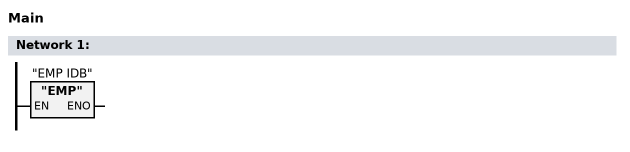
   RUNG wire#powerrail
      "EMP IDB"()
   END_RUNG
   // the same network as SCL:
   "EMP IDB"();   // "EMP"
END_REGION
END_ORGANIZATION_BLOCK

// folder: Display: LED

FUNCTION_BLOCK "LED_Request_Table"   // FB60, SCL
{ S7_Optimized_Access := 'TRUE' }
VERSION : 0.1
   VAR_INPUT
      pn_library : "Recipe: PN Text Library";
      saved_wips : "Recipe: HMI Stations Saved Wips";
      stations : "Station: All Stations";
      table_data : "Part Request Data";
   END_VAR
   VAR_IN_OUT
      request_table : "LED Sign Data";
   END_VAR
   VAR
      row_indices : Array[0..11] of DInt;
   END_VAR
   // row_indices[0] := 0;
   // row_indices[1] := 1;
   // row_indices[2] := 2;
   // row_indices[3] := 3;
   // row_indices[4] := 4;
   // row_indices[5] := 5;
   // row_indices[6] := 6;
   // row_indices[7] := 7;
   // row_indices[8] := 8;
   // row_indices[9] := 9;
   // row_indices[10] := 10;
   // row_indices[11] := 11;
BEGIN
   "Request_Table.Draw"(pn_library := #pn_library,
                        row_indices := #row_indices,
                        saved_wips := #saved_wips,
                        stations := #stations,
                        table_data := #table_data,
                        request_table := #request_table.row);
END_FUNCTION_BLOCK

// folder: Display: Warehouse/001 Request Table

FUNCTION_BLOCK "HMI_Request_Table"   // FB16, SCL
{ S7_Optimized_Access := 'TRUE' }
VERSION : 0.1
   VAR_INPUT
      pn_library : "Recipe: PN Text Library";
      saved_wips : "Recipe: HMI Stations Saved Wips";
      stations : "Station: All Stations";
      table_data : "Part Request Data";
   END_VAR
   VAR_IN_OUT
      barcode_data : "Barcode.UDT";
      request_table : "Part Call Screen";
      request_table_navigation : "Nav Bar Data: PLC";
   END_VAR
   VAR RETAIN
      row_indices : Array[0.."PART_REQUEST_ROW_COUNT_WAREHOUSE_HMI"] of DInt;
   END_VAR
   VAR
      Table_Navigation : "Table Nav";
      Row_Selection : "Request_Table.Row_Selection";
   END_VAR
   // row_indices[1] := 1;
   // row_indices[2] := 2;
   // row_indices[3] := 3;
   // row_indices[4] := 4;
   // row_indices[5] := 5;
   // row_indices[6] := 6;
   // row_indices[7] := 7;
   // row_indices[8] := 8;
   // row_indices[9] := 9;
   // row_indices[10] := 10;
BEGIN
   REGION "TABLE NAVIGATION"
       #Table_Navigation(tblData := #table_data.row,
                         tblDisp := #request_table.row,
                         tableNav := #request_table_navigation,
                         rowIndices := #row_indices);
   END_REGION


   REGION "NAV BUTTON ANIMATIONS"
       "Request_Table.Navigation_Animations"(#request_table_navigation);
   END_REGION


   REGION "DRAW TABLE"
       "Request_Table.Draw"(pn_library := #pn_library,
                            row_indices := #row_indices,
                            saved_wips := #saved_wips,
                            stations := #stations,
                            table_data := #table_data,
                            request_table := #request_table.row);
   END_REGION


   REGION "LOAD SELECTION DATA"
       #Row_Selection(request_table := #request_table,
                      barcode_data := #barcode_data);
   END_REGION
END_FUNCTION_BLOCK

FUNCTION "Address in Loaded Wip" : Bool   // FC43, SCL
{ S7_Optimized_Access := 'TRUE' }
VERSION : 0.1
   VAR_INPUT
      pWip : DInt;
      stn : "Station: Single Station";
   END_VAR
   VAR_TEMP
      ret : Bool;
   END_VAR
BEGIN
   IF #pWip = #stn.wipData.index THEN
       #ret := TRUE;
   END_IF;
   #"Address in Loaded Wip" := #ret;
END_FUNCTION

// folder: Display: Warehouse/002 Settings

FUNCTION_BLOCK "Settings Screen"   // FB19, SCL
{ S7_Optimized_Access := 'TRUE' }
VERSION : 0.1
   VAR_INPUT
      settings_meta : "Setting Meta Data";
      wip_library : "Recipe: Wip Text Library";
   END_VAR
   VAR_IN_OUT
      pn_library : "Recipe: PN Text Library";
      saved_wips : "Recipe: HMI Stations Saved Wips";
      stations : "Station: All Stations";
      settings : "Settings";
   END_VAR
   VAR
      "Assign Button" : "Assign Button";
      "Critical Time IO Field" : "Critical_IO_Field";
      "Dropzone IO Field" : "Dropzone_IO_Field";
      first_row : DInt;
      "Line IO Field" : "Line_IO_Field";
      "Part Number IO Field" : "Part Number IO Field";
      processed_inputs : "Settings Screen: Processed Inputs";
      "Select Buttons Button" : "Select Buttons";
      "Select Station Button" : "Select Station PB";
      "Select WIP Button" : "Select WIP PB";
      "Table Nav_Instance" : "Table Nav";
      "Total Time IO Field" : "Total_IO_Field";
      "WIP Select Table NavBar" : "NavBar";
      inst_Selected_WIP_Table : "Selected_WIP_Table";
   END_VAR
   VAR_TEMP
      _station_rows_buffer : Array[0..2] of "Settings Station Row Data";
   END_VAR
   VAR CONSTANT
      TABLE_LENGTH : DInt := 49;
      VISIBLE_ROW_COUNT : DInt := 2;
   END_VAR
BEGIN
   REGION "SELECT STATION BUTTON"
       #"Select Station Button"(#settings.selectStation);
   END_REGION

   REGION "SELECT BUTTONS BUTTON"
       #"Select Buttons Button"(settings_meta := #settings_meta,
                                stations := #stations,
                                interface := #settings.selectButton);
   END_REGION

   REGION "SELECT WIP BUTTON"
       #"Select WIP Button"(settings_meta := #settings_meta,
                            stations := #stations,
                            interface := #settings.selectWip);
   END_REGION

   REGION "LINE IO FIELD"
       #"Line IO Field"(settings_meta := #settings_meta,
                        stations := #stations,
                        interface := #settings.line,
                        get_line := #processed_inputs.line_name);
   END_REGION

   REGION "DROPZONE IO FIELD"
       #"Dropzone IO Field"(settings_meta := #settings_meta,
                            stations := #stations,
                            interface := #settings.dropzone,
                            get_dropzone := #processed_inputs.dropzone);
   END_REGION

   REGION "TOTAL TIME IO FIELD"
       #"Total Time IO Field"(settings_meta := #settings_meta,
                              stations := #stations,
                              interface := #settings.total,
                              state_changes := #processed_inputs.total);
   END_REGION

   REGION "CRITICAL TIME IO FIELD"
       #"Critical Time IO Field"(settings_meta := #settings_meta,
                                 stations := #stations,
                                 interface := #settings.critical,
                                 state_changes := #processed_inputs.critical);
   END_REGION

   REGION "PART NUMBER ENTRY FIELD"
       #"Part Number IO Field"(settings_meta := #settings_meta,
                               stations := #stations,
                               part_number_library := #pn_library,
                               interface := #settings.partNumber,
                               processed_part_number_entry := #processed_inputs.part_number);

   END_REGION

   REGION "ASSIGN BUTTON"
       #"Assign Button"(processed_inputs := #processed_inputs,
                        settings := #settings,
                        settings_meta := #settings_meta,
                        pn_library := #pn_library,
                        saved_wips := #saved_wips,
                        stations := #stations,
                        interface := #settings.assign,
                        state_changes := #processed_inputs.assign);
   END_REGION

   REGION "SELECTED WIP TABLE"
       #_station_rows_buffer := #settings.stationRows;
       #inst_Selected_WIP_Table(saved_wips := #saved_wips,
                                settings_meta := #settings_meta,
                                stations := #stations,
                                wip_library := #wip_library,
                                pn_library := #pn_library,
                                navigation_bar := #settings.stnTableNavBar.plc,
                                stationRows := #_station_rows_buffer);
       #settings.stationRows := #_station_rows_buffer;
   END_REGION

   REGION "WIP SELECT TABLE NAVBAR"
       #"WIP Select Table NavBar"(hide := #settings_meta.selected_stations.count < 4,
                                  TABLE_LENGTH := #TABLE_LENGTH,
                                  VISIBLE_ROW_COUNT := #VISIBLE_ROW_COUNT,
                                  interface := #settings.stnTableNavBar,
                                  first_row := #first_row);
   END_REGION
END_FUNCTION_BLOCK

FUNCTION "Settings Screen: Load Selected: Non-HMI Station" : Void   // FC150, SCL
{ S7_Optimized_Access := 'TRUE' }
VERSION : 0.1
   VAR_INPUT
      stations : "Station: All Stations";
      selected_stations : "Selected Stations";
      wip_library : "Recipe: Wip Text Library";
      part_number_library : "Recipe: PN Text Library";
   END_VAR
   VAR_IN_OUT
      selected_station_table : Array[0..2] of "Settings Station Row Data";
   END_VAR
   VAR_TEMP
      station_index : Int;
      table_row_index : Int;
   END_VAR
BEGIN
   FOR #station_index := 0 TO "STATION_COUNT" DO
       IF #selected_stations.stns[#station_index] THEN
           "Settings Screen: Load Selected WIP"(station := #stations.stn[#station_index],
                                                wip_library := #wip_library,
                                                part_number_library := #part_number_library,
                                                table_row := #selected_station_table[#table_row_index]);
           #table_row_index += 1;
           IF #table_row_index > 2 THEN
               EXIT;
           END_IF;
       END_IF;
   END_FOR;
END_FUNCTION

FUNCTION "Settings Screen: Load Selected WIP" : Void   // FC151, SCL
{ S7_Optimized_Access := 'TRUE' }
VERSION : 0.1
   VAR_INPUT
      station : "Station: Single Station";
      wip_library : "Recipe: Wip Text Library";
      part_number_library : "Recipe: PN Text Library";
   END_VAR
   VAR_IN_OUT
      table_row : "Settings Station Row Data";
   END_VAR
   VAR_TEMP
      _table_row : "Settings Station Row Data";
      button_index : Int;
   END_VAR
BEGIN
   REGION "NOTES"
       (*
       Simple data map from station presented at input to hmi data structure.
       Decision about which data to map is done in parent.
       last edit: 2021-10-06
       *)
   END_REGION

   REGION "BUFFER IN"
       #_table_row := #table_row;
   END_REGION

   REGION "MAP"
       #_table_row.line.data := #station.id.lineName;
       #_table_row.dropzone.data := "Strip Sign"(USINT_TO_WSTRING(#station.id.dropZone));
       #_table_row.wip.data := "WIP.Code_to_WString"(wipTxtLib := #wip_library,
                                                           code := #station.wipData.code);
       FOR #button_index := 0 TO "BUTTON_COUNT" DO
           "Settings Screen: Load Selected WIP: Load Button"(wip_components:=#station.wipCmpts,
                                                                 wip_library := #wip_library,
                                                                 button_index := #button_index,
                                                                 part_number_liberary := #part_number_library,
                                                                 button_row := #_table_row.btnRows[#button_index]);
       END_FOR;
   END_REGION

   REGION "BUFFER OUT"
       #table_row := #_table_row;
   END_REGION
END_FUNCTION

FUNCTION "Settings Screen: Selected Station Table Row Color" : Void   // FC152, SCL
{ S7_Optimized_Access := 'TRUE' }
VERSION : 0.1
BEGIN
END_FUNCTION

FUNCTION "Settings Screen: Load Selected WIP: Load Button" : Void   // FC155, SCL
{ S7_Optimized_Access := 'TRUE' }
VERSION : 0.1
   VAR_INPUT
      button_index : Int;
      part_number_liberary : "Recipe: PN Text Library";
      wip_components : "Station: Wip: Wip Module";
      wip_library : "Recipe: Wip Text Library";
   END_VAR
   VAR_IN_OUT
      button_row : "Settings Station Row Button Row Data";
   END_VAR
   VAR_TEMP
      _button_row : "Settings Station Row Button Row Data";
      part_number_wstring : WString;
      part_number_code : DInt;
   END_VAR
   VAR CONSTANT
      no_code : WString;
   END_VAR
BEGIN
   REGION "NOTES"
       (*
       Simple data map from station presented at input to hmi data structure.
       Decision about which data to map is done in parent.
       last edit: 2021-10-06
       *)
   END_REGION

   REGION "BUFFER IN"    
       #_button_row := #button_row;
   END_REGION

   REGION "BUTTON LABEL"
       // CURRENTLY A STATIC LABEL
   END_REGION

   REGION "ALOTTED TIME"
       #_button_row.total.data := "Timer.Real_to_WString"(#wip_components.timers.ptAllotted[#button_index]);
   END_REGION

   REGION "CRITICAL TIME"
       #_button_row.critical.data := "Timer.Real_to_WString"(#wip_components.timers.ptCritical[#button_index]);
   END_REGION

   REGION "PART NUMBER"

       REGION "PROCESS PART NUMBER"
           #part_number_code := #wip_components.pnCode[#button_index];
           #part_number_wstring := "Part_Number.Code_to_WString"(pnLib := #part_number_liberary,
                                                         pnCode := #part_number_code);
       END_REGION

       REGION "SINGLE LINE PART NUMBER"
           IF "Part_Number.Is_Single"(#part_number_code) THEN
               #_button_row.singlePN.data := #part_number_wstring;
               #_button_row.doublePN.data := #no_code;
           END_IF;
       END_REGION

       REGION "DOUBLE LINE PART NUMBER"
           IF "Part_Number.Is_Double"(#part_number_code) THEN
               #_button_row.singlePN.data := #no_code;
               #_button_row.doublePN.data := #part_number_wstring;
           END_IF;
       END_REGION

   END_REGION

   REGION "BUFFER OUT"
       #button_row := #_button_row;
   END_REGION
END_FUNCTION

FUNCTION "Settings Screen: Load Selected: HMI Station" : Void   // FC176, SCL
{ S7_Optimized_Access := 'TRUE' }
VERSION : 0.1
   VAR_INPUT
      stations : "Station: All Stations";
      selected_wips : "Selected Wips";
      wip_library : "Recipe: Wip Text Library";
      part_number_library : "Recipe: PN Text Library";
   END_VAR
   VAR_IN_OUT
      selected_station_table : Array[0..2] of "Settings Station Row Data";
   END_VAR
   VAR_TEMP
      station_index : Int;
      table_row_index : Int;
   END_VAR
BEGIN
   FOR #station_index := 0 TO #selected_wips.count DO
       "Settings Screen: Load Selected WIP"(station := #stations.stn[#station_index],
                                            wip_library := #wip_library,
                                            part_number_library := #part_number_library,
                                            table_row := #selected_station_table[#table_row_index]);END_FOR;
END_FUNCTION

// folder: Display: Warehouse/002 Settings/Assign Button

FUNCTION_BLOCK "Assign Button"   // FB55, SCL
{ S7_Optimized_Access := 'TRUE' }
VERSION : 0.1
   VAR_INPUT
      processed_inputs : "Settings Screen: Processed Inputs";
      settings : "Settings";
      settings_meta : "Setting Meta Data";
   END_VAR
   VAR_IN_OUT
      interface : "Push Button Data";
      pn_library : "Recipe: PN Text Library";
      saved_wips : "Recipe: HMI Stations Saved Wips";
      state_changes : "Push Button Data: State Change Data";
      stations : "Station: All Stations";
   END_VAR
   VAR
      "Push Button: State Changes" : "Push Button: State Changes";
   END_VAR
   VAR_TEMP
      _interface : "Push Button Data";
      _state_changes : "Push Button Data: State Change Data";
   END_VAR
BEGIN
   REGION "BUFFER IN"
       #_interface := #interface;
   END_REGION


   REGION "PROCESS USER INPUT"
       #"Push Button: State Changes"(interface := #_interface,
                                     state_changes := #_state_changes);
   END_REGION


   REGION "ANIMATE"
       "Assign_Button.Animate"(settings_meta := #settings_meta,
                                         interface := #_interface);
   END_REGION


   REGION "PERFOM ASSIGNMNET"
       IF #_state_changes.actuate.falling THEN
           "Assign_Button.Perform_Assignment"(processed_inputs := #processed_inputs,
                                              settings := #settings,
                                              settings_meta := #settings_meta,
                                              pn_library := #pn_library,
                                              stations := #stations,
                                              saved_wips := #saved_wips);
       END_IF;
   END_REGION


   REGION "BUFFER OUT"
       #interface := #_interface;
       #state_changes := #_state_changes;
   END_REGION
END_FUNCTION_BLOCK

FUNCTION "Assign_Button.Make_Visible_Enable" : Bool   // FC197, SCL
{ S7_Optimized_Access := 'TRUE' }
VERSION : 0.1
   VAR_INPUT
      setting_meta : "Setting Meta Data";
   END_VAR
BEGIN
   #"Assign_Button.Make_Visible_Enable" :=  #setting_meta.selected_btns.count > 0;
END_FUNCTION

FUNCTION "Assign_Button.Animate" : Void   // FC198, SCL
{ S7_Optimized_Access := 'TRUE' }
VERSION : 0.1
   VAR_INPUT
      settings_meta : "Setting Meta Data";
   END_VAR
   VAR_IN_OUT
      interface : "Push Button Data";
   END_VAR
   VAR_TEMP
      selected_station_count : DInt;
   END_VAR
BEGIN
   REGION "COLOR"
   #interface.animate := "WHITE_BACKGROUND";
   END_REGION

   REGION "VISIBILITY
       #interface.visible := "Assign_Button.Make_Visible_Enable"(setting_meta := #settings_meta);
   END_REGION

   REGION "ENABLE"
       #interface.enable := "Assign_Button.Make_Visible_Enable"(setting_meta := #settings_meta);
   END_REGION
END_FUNCTION

FUNCTION "Assign_Button.Perform_Assignment" : Void   // FC235, SCL
{ S7_Optimized_Access := 'TRUE' }
VERSION : 0.1
   VAR_INPUT
      processed_inputs : "Settings Screen: Processed Inputs";
      settings : "Settings";
      settings_meta : "Setting Meta Data";
   END_VAR
   VAR_IN_OUT
      pn_library : "Recipe: PN Text Library";
      stations : "Station: All Stations";
      saved_wips : "Recipe: HMI Stations Saved Wips";
   END_VAR
   VAR_TEMP
      _station_indices : Array[0.."STATION_COUNT"] of Int;
   END_VAR
BEGIN
   REGION "DO NOTHING ON NO SELECTED STAION"
       IF #settings_meta.selected_stations.count = 0 THEN
           RETURN;
       END_IF;
   END_REGION


   REGION "HMI STATIONS"
       "Selected_Stations.Indices"(selected_stations:=#settings_meta.selected_stations,
                                   selected_stations_indices:=#_station_indices);
       IF "Is_HMI_Station"(#stations.stn[#_station_indices[0]]) THEN
           "Assign_Button.HMI_Stations"(processed_inputs := #processed_inputs,
                                        settings := #settings,
                                        settings_meta := #settings_meta,
                                        pn_library := #pn_library,
                                        saved_wips := #saved_wips,
                                        stations := #stations);
           RETURN;
       END_IF;
   END_REGION


   REGION "KP8 STATIONS"
       "Assign_Button.KP8_Station"(processed_inputs := #processed_inputs,
                                   settings := #settings,
                                   settings_meta := #settings_meta,
                                   all_stations := #stations,
                                   pn_library := #pn_library);
       RETURN;
   END_REGION
END_FUNCTION

FUNCTION "Assign_Button.Assign_ID_Parameters" : Void   // FC264, SCL
{ S7_Optimized_Access := 'TRUE' }
VERSION : 0.1
   VAR_INPUT
      processed_inputs : "Settings Screen: Processed Inputs";
      settings : "Settings";
   END_VAR
   VAR_IN_OUT
      id : "Station: Id";
   END_VAR
BEGIN
   IF #settings.line.enable THEN
       #id.lineName := #processed_inputs.line_name.actual;
   END_IF;
   IF #settings.dropzone.enable THEN
       #id.dropZone := #processed_inputs.dropzone.actual;
   END_IF;
END_FUNCTION

// folder: Display: Warehouse/002 Settings/Assign Button/HMI Station

FUNCTION "Assign_Button.HMI_Stations" : Void   // FC236, SCL
{ S7_Optimized_Access := 'TRUE' }
VERSION : 0.1
   VAR_INPUT
      processed_inputs : "Settings Screen: Processed Inputs";
      settings : "Settings";
      settings_meta : "Setting Meta Data";
   END_VAR
   VAR_IN_OUT
      pn_library : "Recipe: PN Text Library";
      saved_wips : "Recipe: HMI Stations Saved Wips";
      stations : "Station: All Stations";
   END_VAR
   VAR_TEMP
      _i : Int;
      _length : Int;
      _selected_stations : Array[0.."STATION_COUNT"] of Int;
      _p_station : Int;
   END_VAR
BEGIN
   REGION "DO NOTHING IF NO STATIONS SELECTED"
       IF #settings_meta.selected_stations.count = 0 THEN
           RETURN;
       END_IF;
   END_REGION


   REGION "GET INDICES OF SELECTED STATIONS"
       "Selected_Stations.Indices"(selected_stations := #settings_meta.selected_stations,
                                   selected_stations_indices := #_selected_stations);

   END_REGION


   REGION "FOR EACH SELECTED STATION"
       #_length := UDINT_TO_INT("Array.Any.Length"(#saved_wips.stn)) - 1;
       FOR #_i := 0 TO #_length DO

           IF #_selected_stations[#_i] = "NULL_TOKEN" THEN
               RETURN;
           END_IF;

           REGION "ASSIGN TO WIP"
               "Assign_Button.Assign_ID_Parameters"(processed_inputs := #processed_inputs,
                                                    settings := #settings,
                                                    id := #stations.stn[#_selected_stations[#_i]].id);
               #_p_station := "WIP.Global_Index_to_HMI_Station_Index"(global_index := #_selected_stations[#_i],
                                                                      saved_WIPs := #saved_wips);
               "Assign_Button.HMI_Stations.WIP"(processed_inputs:=#processed_inputs,
                                                selected_wips := #settings_meta.selected_wips,
                                                selected_buttons := #settings_meta.selected_btns,
                                                pn_library := #pn_library,
                                                stations_wips := #saved_wips.stn[#_p_station]);
           END_REGION

       END_FOR;
   END_REGION
END_FUNCTION

FUNCTION "Assign_Button.HMI_Stations.WIP" : Void   // FC237, SCL
{ S7_Optimized_Access := 'TRUE' }
VERSION : 0.1
   VAR_INPUT
      processed_inputs : "Settings Screen: Processed Inputs";
      selected_wips : "Selected Wips";
      selected_buttons : "Selected Buttons";
   END_VAR
   VAR_IN_OUT
      pn_library : "Recipe: PN Text Library";
      stations_wips : "WIP: Station";
   END_VAR
   VAR_TEMP
      _i : Int;
      _p_wip : Int;
      _selected_wip_indices : Array[0.."WIP_COUNT"] of Int;
   END_VAR
BEGIN
   REGION "DO NOTHING IF NO WIPS SELECTED"
       IF #selected_wips.count = 0 THEN
           RETURN;
       END_IF;
   END_REGION


   REGION "GET INDICES OF SELECTED WIPS"    
       "WIP_Station.Indices_of_Selected_WIPs"(selected_wips := #selected_wips,
                                              station_wips := #stations_wips,
                                              selected_wip_indices := #_selected_wip_indices);
   END_REGION


   REGION "FOR EACH SELECTED WIP"
       FOR #_i := 0 TO #selected_wips.count DO

           REGION "ASSIGN DATA TO SELECTED BUTTONS"
               #_p_wip := #_selected_wip_indices[#_i];
               IF #_p_wip = "NULL_TOKEN" THEN
                   RETURN;
               END_IF;
               "Assign_Button.HMI_Stations.WIP.Buttons"(processed_inputs := #processed_inputs,
                                                        selected_buttons := #selected_buttons,
                                                        pn_library := #pn_library,
                                                        wip_module := #stations_wips.wip[#_p_wip]);
           END_REGION

       END_FOR;
   END_REGION
END_FUNCTION

FUNCTION "Assign_Button.HMI_Stations.WIP.Buttons" : Void   // FC238, SCL
{ S7_Optimized_Access := 'TRUE' }
VERSION : 0.1
   VAR_INPUT
      processed_inputs : "Settings Screen: Processed Inputs";
      selected_buttons : "Selected Buttons";
   END_VAR
   VAR_IN_OUT
      pn_library : "Recipe: PN Text Library";
      wip_module : "Station: Wip: Wip Module";
   END_VAR
   VAR_TEMP
      _i : Int;
      _p_btn : Int;
      _selected_buttons_indices : Array[0..7] of Int;
   END_VAR
BEGIN
   REGION "DO NOTHING IF NO BUTTONS SELECTED
       IF #selected_buttons.count = 0 THEN
           RETURN;
       END_IF;
   END_REGION


   REGION "GET INDICES OF SELECTED BUTTONS"
       "Selected_Buttons.Indices"(selected_buttons := #selected_buttons,
                                  selected_buttons_indices := #_selected_buttons_indices);
   END_REGION

   REGION "FOR EACH SELECTED BUTTON"
       FOR #_i := 0 TO #selected_buttons.count DO

           REGION "ASSIGN DATA TO SELECTED BUTTON"
               #_p_btn := #_selected_buttons_indices[#_i];
               "Assign_Button.HMI_Stations.Assign_Station_Button_Data"(processed_inputs := #processed_inputs,
                                                                       index := #_p_btn,
                                                                       pn_library := #pn_library,
                                                                       wip_module := #wip_module);
           END_REGION

       END_FOR;
   END_REGION
END_FUNCTION

FUNCTION "Assign_Button.HMI_Stations.Assign_Station_Button_Data" : Void   // FC239, SCL
{ S7_Optimized_Access := 'TRUE' }
VERSION : 0.1
   VAR_INPUT
      processed_inputs : "Settings Screen: Processed Inputs";
      index : Int;
   END_VAR
   VAR_IN_OUT
      pn_library : "Recipe: PN Text Library";
      wip_module : "Station: Wip: Wip Module";
   END_VAR
BEGIN
   IF #index = "NULL_TOKEN" THEN
       RETURN;
   END_IF;
   #wip_module.pnCode[#index] := "Part_Number.WString_to_Code"(part_number := #processed_inputs.part_number.actual,
                                                               pn_library := #pn_library);
   #wip_module.timers.ptAllotted[#index] := #processed_inputs.total.actual;
   #wip_module.timers.ptCritical[#index] := #processed_inputs.critical.actual;
END_FUNCTION

// folder: Display: Warehouse/002 Settings/Assign Button/KP8 Station

FUNCTION "Assign_Button.KP8_Station" : Void   // FC247, SCL
{ S7_Optimized_Access := 'TRUE' }
VERSION : 0.1
   VAR_INPUT
      processed_inputs : "Settings Screen: Processed Inputs";
      settings : "Settings";
      settings_meta : "Setting Meta Data";
   END_VAR
   VAR_IN_OUT
      all_stations : "Station: All Stations";
      pn_library : "Recipe: PN Text Library";
   END_VAR
   VAR_TEMP
      _i : Int;
      _length : Int;
      _selected_stations : Array[0.."STATION_COUNT"] of Int;
      _p_station : Int;
   END_VAR
BEGIN
   REGION "DO NOTHING IF NO STATIONS SELECTED"
       IF #settings_meta.selected_stations.count = 0 THEN
           RETURN;
       END_IF;
   END_REGION


   REGION "GET INDICES OF SELECTED STATIONS"
       "Selected_Stations.Indices"(selected_stations := #settings_meta.selected_stations,
                                   selected_stations_indices := #_selected_stations);
   END_REGION


   REGION "FOR EACH SELECTED STATION"
       IF #settings_meta.selectable_stations.count = 0 THEN
           RETURN;
       END_IF;
       FOR #_i := 0 TO #settings_meta.selected_stations.count DO
           IF #_selected_stations[#_i] = "NULL_TOKEN" THEN
               RETURN;
           END_IF;
           #_p_station := #_selected_stations[#_i];
           "Assign_Button.Assign_ID_Parameters"(processed_inputs := #processed_inputs,
                                                settings := #settings,
                                                id := #all_stations.stn[#_p_station].id);
           "Assign_Button.KP8_Stations.Buttons"(processed_inputs := #processed_inputs,
                                                selected_buttons := #settings_meta.selected_btns,
                                                pn_library := #pn_library,
                                                station := #all_stations.stn[#_p_station]);
       END_FOR;
   END_REGION
END_FUNCTION

FUNCTION "Assign_Button.KP8_Station.Assign_Station_Button_Data" : Void   // FC248, SCL
{ S7_Optimized_Access := 'TRUE' }
VERSION : 0.1
   VAR_INPUT
      button_number : Int;
      processed_inputs : "Settings Screen: Processed Inputs";
   END_VAR
   VAR_IN_OUT
      pn_library : "Recipe: PN Text Library";
      station : "Station: Single Station";
   END_VAR
   VAR_TEMP
      _i : Int;
      _length : Int;
      _selected_stations : Array[0.."STATION_COUNT"] of Int;
      _p_station : Int;
   END_VAR
BEGIN
   IF #button_number = "NULL_TOKEN" THEN
       RETURN;
   END_IF;
   #station.wipCmpts.pnCode[#button_number] := "Part_Number.WString_to_Code"(part_number := #processed_inputs.part_number.actual,
                                                                             pn_library := #pn_library);
   #station.wipCmpts.timers.ptCritical[#button_number] := #processed_inputs.critical.actual;
   #station.wipCmpts.timers.ptAllotted[#button_number] := #processed_inputs.total.actual;
END_FUNCTION

FUNCTION "Assign_Button.KP8_Stations.Buttons" : Void   // FC249, SCL
{ S7_Optimized_Access := 'TRUE' }
VERSION : 0.1
   VAR_INPUT
      processed_inputs : "Settings Screen: Processed Inputs";
      selected_buttons : "Selected Buttons";
   END_VAR
   VAR_IN_OUT
      pn_library : "Recipe: PN Text Library";
      station : "Station: Single Station";
   END_VAR
   VAR_TEMP
      _i : Int;
      _p_btn : Int;
      _selected_buttons_indices : Array[0..7] of Int;
   END_VAR
BEGIN
   REGION "DO NOTHING IF NO BUTTONS SELECTED
       IF #selected_buttons.count = 0 THEN
           RETURN;
       END_IF;
   END_REGION


   REGION "GET INDICES OF SELECTED BUTTONS"
       "Selected_Buttons.Indices"(selected_buttons := #selected_buttons,
                                  selected_buttons_indices := #_selected_buttons_indices);
   END_REGION


   REGION "FOR EACH SELECTED BUTTON"
       FOR #_i := 0 TO #selected_buttons.count - 1 DO

           IF #_selected_buttons_indices[#_i] = "NULL_TOKEN" THEN
               RETURN;
           END_IF;

           REGION "ASSIGN DATA TO SELECTED BUTTON"
               #_p_btn := #_selected_buttons_indices[#_i];
               "Assign_Button.KP8_Station.Assign_Station_Button_Data"(button_number := #_p_btn,
                                                                      processed_inputs := #processed_inputs,
                                                                      pn_library := #pn_library,
                                                                      station := #station);
           END_REGION

       END_FOR;
   END_REGION
END_FUNCTION

// folder: Display: Warehouse/002 Settings/Critical IO Field

FUNCTION_BLOCK "Critical_IO_Field"   // FB53, SCL
{ S7_Optimized_Access := 'TRUE' }
VERSION : 0.1
   VAR_INPUT
      settings_meta : "Setting Meta Data";
      stations : "Station: All Stations";
   END_VAR
   VAR_IN_OUT
      interface : "IO Field Data: Label with Data";
      state_changes : "State Changes: Real";
   END_VAR
   VAR
      Critical_IO_Field : "IO Field: State Changes";
      Detect_Stat_Changes : "Real.State_Change";
   END_VAR
   VAR_TEMP
      _interface : "IO Field Data: Label with Data";
      feedback : "IO Field: State Change Data";
   END_VAR
BEGIN
   REGION "BUFFER IN"
       #_interface := #interface;
   END_REGION

   REGION "PROCESS USER INPUT"
       #Critical_IO_Field(interface := #_interface,
                          feedback := #feedback);
       #Detect_Stat_Changes(value := "Timer.WString_to_Real"(#_interface.value),
                            get_real := #state_changes);
   END_REGION

   REGION "BUFFER OUT"
       "Critical_IO_Field.Animate"(feedback := #feedback,
                                   settings_meta := #settings_meta,
                                   stations := #stations,
                                   interface := #_interface);
   END_REGION

   REGION "BUFFER OUT"
       #interface := #_interface;
   END_REGION
END_FUNCTION_BLOCK

FUNCTION "Critical_IO_Field.Make_Visible_Enable" : Bool   // FC191, SCL
{ S7_Optimized_Access := 'TRUE' }
VERSION : 0.1
   VAR_INPUT
      setting_meta : "Setting Meta Data";
   END_VAR
BEGIN
   #"Critical_IO_Field.Make_Visible_Enable" :=  #setting_meta.selected_btns.count > 0;
END_FUNCTION

FUNCTION "Critical_IO_Field.Animate" : Void   // FC192, SCL
{ S7_Optimized_Access := 'TRUE' }
VERSION : 0.1
   VAR_INPUT
      feedback : "IO Field: State Change Data";
      settings_meta : "Setting Meta Data";
      stations : "Station: All Stations";
   END_VAR
   VAR_IN_OUT
      interface : "IO Field Data: Label with Data";
   END_VAR
   VAR_TEMP
      _visible_enabled : Bool;
   END_VAR
BEGIN
   REGION "COLOR"
   #interface.animate := "WHITE_BACKGROUND";
   END_REGION


   REGION "SET STATE"
       #_visible_enabled := "Critical_IO_Field.Make_Visible_Enable"(setting_meta := #settings_meta);
   END_REGION


   REGION "VISIBILITY
       #interface.visible := #_visible_enabled;
   END_REGION


   REGION "ENABLE"
       #interface.enable := #_visible_enabled;
   END_REGION


   REGION "POPULATE VALUE"
       IF #settings_meta.button_selection_change.selection_change THEN
           #interface.value := "Critical_IO_Field.Populate_Value"(hidden := NOT #_visible_enabled,
                                                                  selected_buttons := #settings_meta.selected_btns,
                                                                  selected_stations := #settings_meta.selected_stations,
                                                                  stations := #stations);
       END_IF;
   END_REGION
END_FUNCTION

FUNCTION "Critical_IO_Field.Populate_Value" : WString   // FC283, SCL
{ S7_Optimized_Access := 'TRUE' }
VERSION : 0.1
   VAR_INPUT
      hidden : Bool;
      selected_buttons : "Selected Buttons";
      selected_stations : "Selected Stations";
      stations : "Station: All Stations";
   END_VAR
   VAR_TEMP
      _critical : WString;
      _p_station : Int;
      _p_button : Int;
   END_VAR
   VAR CONSTANT
      BLANK : WString;
      ZERO : WChar := WCHAR#'0';
   END_VAR
BEGIN
   IF #hidden THEN
       #"Critical_IO_Field.Populate_Value" := #BLANK;
       RETURN;
   END_IF;
   #_p_station := "Selected_Stations.Get_First_Selected_Station"(#selected_stations);
   #_p_button := "Selected_Buttons.Get_First_Selected_Button"(#selected_buttons);
   #_critical := "Timer.Real_to_WString"(#stations.stn[#_p_station].wipCmpts.timers.ptCritical[#_p_button]);
   #"Critical_IO_Field.Populate_Value" := #_critical;
END_FUNCTION

// folder: Display: Warehouse/002 Settings/Dropzone IO Field

FUNCTION_BLOCK "Dropzone_IO_Field"   // FB50, SCL
{ S7_Optimized_Access := 'TRUE' }
VERSION : 0.1
   VAR_INPUT
      settings_meta : "Setting Meta Data";
      stations : "Station: All Stations";
   END_VAR
   VAR_IN_OUT
      interface : "IO Field Data: Label with Data";
      get_dropzone : "State Changes: USInt";
   END_VAR
   VAR
      "Line IO Field" : "IO Field: State Changes";
      "Get Dropzone Input" : "USInt.State_change";
   END_VAR
   VAR_TEMP
      _feedback : "IO Field: State Change Data";
      _interface : "IO Field Data: Label with Data";
   END_VAR
BEGIN
   REGION "BUFFER IN"
       #_interface := #interface;
   END_REGION


   REGION "PROCESS USER INPUT"
       #"Line IO Field"(interface := #_interface,
                        feedback := #_feedback);
       #"Get Dropzone Input"(value := WSTRING_TO_USINT(#interface.value),
                             get_usint := #get_dropzone);
   END_REGION


   REGION "ANIMATION"
       "Dropzone_IO_Field.Animate"(feedback := #_feedback,
                                   selected_stations := #settings_meta.selected_stations,
                                   settings_meta := #settings_meta,
                                   stations := #stations,
                                   interface := #_interface);
   END_REGION


   REGION "BUFFER OUT"
       #interface := #_interface;
   END_REGION
END_FUNCTION_BLOCK

FUNCTION "Dropzone_IO_Field.Make Visible_Enable" : Bool   // FC185, SCL
{ S7_Optimized_Access := 'TRUE' }
VERSION : 0.1
   VAR_INPUT
      setting_meta : "Setting Meta Data";
      stations : "Station: All Stations";
   END_VAR
   VAR_TEMP
      first_selected_station : Int;
      ret : Bool;
   END_VAR
BEGIN
   IF #setting_meta.selected_stations.count = 0 THEN
       #"Dropzone_IO_Field.Make Visible_Enable" := FALSE;
       RETURN;
   END_IF;


   IF #setting_meta.selected_stations.count > 1 THEN
       #"Dropzone_IO_Field.Make Visible_Enable" := FALSE;
       RETURN;
   END_IF;


   IF #setting_meta.selected_btns.count = 0 THEN
       #"Dropzone_IO_Field.Make Visible_Enable"  := FALSE;
       RETURN;
   END_IF;


   #"Dropzone_IO_Field.Make Visible_Enable" := TRUE;
END_FUNCTION

FUNCTION "Dropzone_IO_Field.Animate" : Void   // FC186, SCL
{ S7_Optimized_Access := 'TRUE' }
VERSION : 0.1
   VAR_INPUT
      feedback : "IO Field: State Change Data";
      selected_stations : "Selected Stations";
      settings_meta : "Setting Meta Data";
      stations : "Station: All Stations";
   END_VAR
   VAR_IN_OUT
      interface : "IO Field Data: Label with Data";
   END_VAR
   VAR_TEMP
      _visible_enabled : Bool;
   END_VAR
BEGIN
   REGION "COLOR"
       #interface.animate := "WHITE_BACKGROUND";
   END_REGION


   REGION "GET STATE"
       #_visible_enabled := "Dropzone_IO_Field.Make Visible_Enable"(setting_meta := #settings_meta,
                                                                                stations := #stations);
   END_REGION


   REGION "VISIBILITY
       #interface.visible := #_visible_enabled;
   END_REGION


   REGION "ENABLE"
       #interface.enable := #_visible_enabled;
   END_REGION


   REGION "POPULATE VALUE"
       IF #settings_meta.button_selection_change.selection_change THEN
           #interface.value := "Dropzone_IO_Field.Populate_Value"(hidden := NOT #_visible_enabled,
                                                                  selected_stations := #selected_stations,
                                                                  stations := #stations);
       END_IF;
   END_REGION
END_FUNCTION

FUNCTION "Dropzone_IO_Field.Populate_Value" : WString   // FC271, SCL
{ S7_Optimized_Access := 'TRUE' }
VERSION : 0.1
   VAR_INPUT
      hidden : Bool;
      selected_stations : "Selected Stations";
      stations : "Station: All Stations";
   END_VAR
   VAR_TEMP
      _dropzone : WString;
      _p_station : Int;
   END_VAR
   VAR CONSTANT
      BLANK : WString;
      ZERO : WChar := WCHAR#'0';
   END_VAR
BEGIN
   IF #hidden THEN
       #"Dropzone_IO_Field.Populate_Value" := #BLANK;
       RETURN;
   END_IF;
   #_p_station := "Selected_Stations.Get_First_Selected_Station"(#selected_stations);
   #_dropzone := USINT_TO_WSTRING(#stations.stn[#_p_station].id.dropZone);
   #_dropzone := "Strip Sign"(#_dropzone);
   #_dropzone := "Trim"(#_dropzone);
   #_dropzone := "Add Leading"("Leading Character" := #ZERO,
                               "Desired Length" := 2,
                               "String" := #_dropzone);
   #"Dropzone_IO_Field.Populate_Value" := #_dropzone;
END_FUNCTION

// folder: Display: Warehouse/002 Settings/Line IO Field

FUNCTION_BLOCK "Line_IO_Field"   // FB47, SCL
{ S7_Optimized_Access := 'TRUE' }
VERSION : 0.1
   VAR_INPUT
      settings_meta : "Setting Meta Data";
      stations : "Station: All Stations";
   END_VAR
   VAR_IN_OUT
      interface : "IO Field Data: Label with Data";
      get_line : "State Changes: WString";
   END_VAR
   VAR
      "Get Line Value" : "WString.State_Change";
      "Line IO Field" : "IO Field: State Changes";
   END_VAR
   VAR_TEMP
      _interface : "IO Field Data: Label with Data";
      feedback : "IO Field: State Change Data";
   END_VAR
BEGIN
   REGION "BUFFER IN"
       #_interface := #interface;
   END_REGION

   REGION "PROCESS USER INPUT"
       #"Line IO Field"(interface := #_interface,
                        feedback := #feedback);
       #"Get Line Value"(interface := #_interface.value,
                         get_wstring := #get_line);

   END_REGION

   REGION "ANIMATION"
       "Line_IO_Field.Animate"(feedback := #feedback,
                               selected_stations := #settings_meta.selected_stations,
                               settings_meta := #settings_meta,
                               stations := #stations,
                               interface := #_interface);
   END_REGION

   REGION "BUFFER OUT"
       #interface := #_interface;
   END_REGION
END_FUNCTION_BLOCK

FUNCTION "Line_IO_Field.Animate" : Void   // FC124, SCL
{ S7_Optimized_Access := 'TRUE' }
VERSION : 0.1
   VAR_INPUT
      feedback : "IO Field: State Change Data";
      selected_stations : "Selected Stations";
      settings_meta : "Setting Meta Data";
      stations : "Station: All Stations";
   END_VAR
   VAR_IN_OUT
      interface : "IO Field Data: Label with Data";
   END_VAR
   VAR_TEMP
      _visible_and_enabled : Bool;
   END_VAR
BEGIN
   REGION "COLOR"
       #interface.animate := "WHITE_BACKGROUND";
   END_REGION


   REGION "STATE"
       #_visible_and_enabled := "Line_IO_Field.Make_Visible_Enable"(selected_stations:= #selected_stations,
                                                                    setting_meta := #settings_meta,
                                                                    stations := #stations);
   END_REGION


   REGION "VISIBILITY
       #interface.visible := #_visible_and_enabled;
   END_REGION


   REGION "ENABLE"
       #interface.enable := #_visible_and_enabled;
   END_REGION


   REGION "POPULATE VALUE"
       IF #settings_meta.button_selection_change.selection_change THEN
           #interface.value := "Line_IO_Field.Populate_Value"(hidden := NOT #_visible_and_enabled,
                                                              selected_stations := #selected_stations,
                                                              stations := #stations);
       END_IF;
   END_REGION
END_FUNCTION

FUNCTION "Line_IO_Field.Make_Visible_Enable" : Bool   // FC187, SCL
{ S7_Optimized_Access := 'TRUE' }
VERSION : 0.1
   VAR_INPUT
      selected_stations : "Selected Stations";
      setting_meta : "Setting Meta Data";
      stations : "Station: All Stations";
   END_VAR
   VAR_TEMP
      first_selected_station : Int;
      ret : Bool;
   END_VAR
BEGIN
   IF #setting_meta.selected_stations.count = 0 THEN
       #"Line_IO_Field.Make_Visible_Enable" := FALSE;
       RETURN;
   END_IF;

   IF #setting_meta.selected_btns.count = 0 THEN
       #"Line_IO_Field.Make_Visible_Enable" := FALSE;
       RETURN;
   END_IF;

   #"Line_IO_Field.Make_Visible_Enable" := "Selected_Stations.Matching_Line_Names"(stations := #stations,
                                                                                               selected_stations := #selected_stations);
END_FUNCTION

FUNCTION "Line_IO_Field.Populate_Value" : WString   // FC268, SCL
{ S7_Optimized_Access := 'TRUE' }
VERSION : 0.1
   VAR_INPUT
      hidden : Bool;
      selected_stations : "Selected Stations";
      stations : "Station: All Stations";
   END_VAR
   VAR_TEMP
      _p_station : Int;
   END_VAR
   VAR CONSTANT
      BLANK : WString;
   END_VAR
BEGIN
   IF #hidden THEN
       #"Line_IO_Field.Populate_Value" := #BLANK;
       RETURN;
   END_IF;
   #_p_station := "Selected_Stations.Get_First_Selected_Station"(#selected_stations);
   #"Line_IO_Field.Populate_Value" := #stations.stn[#_p_station].id.lineName;
END_FUNCTION

// folder: Display: Warehouse/002 Settings/Part Number IO Field

FUNCTION_BLOCK "Part Number IO Field"   // FB54, SCL
{ S7_Optimized_Access := 'TRUE' }
VERSION : 0.1
   VAR_INPUT
      settings_meta : "Setting Meta Data";
      stations : "Station: All Stations";
      part_number_library : "Recipe: PN Text Library";
   END_VAR
   VAR_IN_OUT
      interface : "Part_Number_Double.UDT";
      processed_part_number_entry : "State Changes: WString";
   END_VAR
   VAR
      Resolve_Feedback : "Part_Number_Double.State_Changes";
      Get_Part_Number : "Part_Number_IO_Field.Get_Part_Number";
      display_mode : String[10] := 'single';
   END_VAR
   VAR_TEMP
      _interface : "Part_Number_Double.UDT";
      feedback : "Part_Number_Double.State_Change.UDT";
   END_VAR
BEGIN
   REGION "BUFFER IN"
       #_interface := #interface;
   END_REGION


   REGION "PROCESS USER INPUT"
       #Resolve_Feedback(interface := #_interface,
                         feedback := #feedback);
       "Part_Number_Double_IO_Field.Set_Mode"(feedback := #feedback,
                                              mode := #display_mode);
       #Get_Part_Number(mode := #display_mode,
                        feedback := #feedback,
                        processed_part_number_entry := #processed_part_number_entry);
   END_REGION


   REGION "ANIMATE"
       "Part_Number_IO_Field.Animate"(display_mode := #display_mode,
                                      settings_meta := #settings_meta,
                                      stations := #stations,
                                      part_number_library := #part_number_library,
                                      interface := #_interface);
   END_REGION


   REGION "BUFFER OUT"
       #interface := #_interface;
   END_REGION
END_FUNCTION_BLOCK

FUNCTION "Part_Number_IO_Field.Make_Visible_Enable" : Bool   // FC195, SCL
{ S7_Optimized_Access := 'TRUE' }
VERSION : 0.1
   VAR_INPUT
      setting_meta : "Setting Meta Data";
      visible_mode : String;
      current_mode : String;
   END_VAR
BEGIN
   IF #setting_meta.selected_btns.count = 0 THEN
       #"Part_Number_IO_Field.Make_Visible_Enable" := FALSE;
       RETURN;
   END_IF;

   #"Part_Number_IO_Field.Make_Visible_Enable" := #visible_mode = #current_mode;
END_FUNCTION

FUNCTION "Part_Number_IO_Field.Animate" : Void   // FC196, SCL
{ S7_Optimized_Access := 'TRUE' }
VERSION : 0.1
   VAR_INPUT
      settings_meta : "Setting Meta Data";
      stations : "Station: All Stations";
      part_number_library : "Recipe: PN Text Library";
   END_VAR
   VAR_IN_OUT
      display_mode : String;
      interface : "Part_Number_Double.UDT";
   END_VAR
   VAR_TEMP
      _double_visible_enabled : Bool;
      _single_visible_enabled : Bool;
   END_VAR
   VAR CONSTANT
      SINGLE : String := 'single';
      DOUBLE : String := 'double';
   END_VAR
BEGIN
   REGION "COLOR"
       #interface.single_animate := "WHITE_BACKGROUND";
       #interface.double_animate := "WHITE_BACKGROUND";
   END_REGION


   REGION "STATE"
       #_single_visible_enabled := "Part_Number_IO_Field.Make_Visible_Enable"(setting_meta := #settings_meta,
                                                                              visible_mode := #SINGLE,
                                                                              current_mode := #display_mode);
       #_double_visible_enabled := "Part_Number_IO_Field.Make_Visible_Enable"(setting_meta := #settings_meta,
                                                                              visible_mode := #DOUBLE,
                                                                              current_mode := #display_mode);
   END_REGION


   REGION "VISIBILITY"
       #interface.single_visible := #_single_visible_enabled;
       #interface.double_visible := #_double_visible_enabled;
   END_REGION


   REGION "ENABLE"
       #interface.single_enable := #interface.single_visible;
       #interface.double_enable := #interface.double_visible;
   END_REGION


   REGION "POPULATE VALUE"
       IF #settings_meta.button_selection_change.selection_change THEN
           "Part_Number_IO_Field.Populate_Value"(stations := #stations,
                                                 settings_meta := #settings_meta,
                                                 part_number_library := #part_number_library,
                                                 display_mode := #display_mode,
                                                 interface := #interface);
       END_IF;
   END_REGION
END_FUNCTION

FUNCTION "Part_Number_IO_Field.Populate_Value" : Void   // FC293, SCL
{ S7_Optimized_Access := 'TRUE' }
VERSION : 0.1
   VAR_INPUT
      part_number_library : "Recipe: PN Text Library";
      stations : "Station: All Stations";
      settings_meta : "Setting Meta Data";
   END_VAR
   VAR_IN_OUT
      display_mode : String;
      interface : "Part_Number_Double.UDT";
   END_VAR
   VAR_TEMP
      _p_button : Int;
      _p_station : Int;
      _part_number_code : DInt;
      _part_number : WString;
      _split_part_numbers : Array[0..1] of WString;
   END_VAR
   VAR CONSTANT
      SINGLE : String := 'single';
      DOUBLE : String := 'double';
   END_VAR
BEGIN
   #_p_button := "Selected_Buttons.Get_First_Selected_Button"(#settings_meta.selected_btns);
   IF #_p_button = "NULL_TOKEN" THEN
       RETURN;
   END_IF;
   #_p_station := "Selected_Stations.Get_First_Selected_Station"(#settings_meta.selected_stations);
   IF #_p_station = "NULL_TOKEN" THEN
       RETURN;
   END_IF;
   #_part_number_code := #stations.stn[#_p_station].wipCmpts.pnCode[#_p_button];
   #_part_number := "Part_Number.Code_to_WString"(pnLib := #part_number_library,
                                                  pnCode := #_part_number_code);
   IF "Part_Number.Is_Single"(#_part_number_code) THEN
       #interface.single_value := #_part_number;
       #display_mode := #SINGLE;
       RETURN;
   END_IF;
   "Part_Number.Split_PNs"(part_number := #_part_number,
                           part_numbers := #_split_part_numbers);
   #interface.double_value_top := #_split_part_numbers[0];
   #interface.double_value_bottom := #_split_part_numbers[1];
   #display_mode := #DOUBLE;
   RETURN;
END_FUNCTION

// folder: Display: Warehouse/002 Settings/Select Buttons Button

FUNCTION_BLOCK "Select Buttons"   // FB42, SCL
{ S7_Optimized_Access := 'TRUE' }
VERSION : 0.1
   VAR_INPUT
      settings_meta : "Setting Meta Data";
      stations : "Station: All Stations";
   END_VAR
   VAR_IN_OUT
      interface : "Push Button Data";
   END_VAR
   VAR
      "Get Button Feedback" : "Push Button: State Changes";
   END_VAR
   VAR_TEMP
      _interface : "Push Button Data";
      enable : Bool;
      feedback : "Push Button Data: State Change Data";
      visible : Bool;
   END_VAR
BEGIN
   REGION "BUFFER IN"
       #_interface := #interface;
   END_REGION

   REGION "PROCESS USER INPUT"
       #"Get Button Feedback"(interface := #_interface,
                              state_changes := #feedback);
   END_REGION

   REGION "ANIMATIONS"
       "Select Buttons: Private: Animations"(feedback := #feedback,
                                             settings_meta := #settings_meta,
                                             stations := #stations,
                                             interface := #_interface);
   END_REGION

   REGION "BUFFER OUT"
       #interface := #_interface;
   END_REGION
END_FUNCTION_BLOCK

FUNCTION "Select Buttons: Private: Animations" : Void   // FC93, SCL
{ S7_Optimized_Access := 'TRUE' }
VERSION : 0.1
   VAR_INPUT
      feedback : "Push Button Data: State Change Data";
      settings_meta : "Setting Meta Data";
      stations : "Station: All Stations";
   END_VAR
   VAR_IN_OUT
      interface : "Push Button Data";
   END_VAR
BEGIN
   REGION "COLOR"
       #interface.animate := "Bool.Animate"(true_color := "GREEN_LIGHT_BACKGROUND",
                                             false_color := "GRAY_BACKGROUND",
                                             evaluation_signal := #feedback.actuate.actual);
   END_REGION

   REGION "VISIBILITY"
       #interface.visible := "Select Buttons: Private: Make Visible / Enable"(settings_meta := #settings_meta,
                                                                               stations := #stations);
   END_REGION

   REGION "ENABLED STATE"
       #interface.enable := "Select Buttons: Private: Make Visible / Enable"(settings_meta := #settings_meta,
                                                                              stations := #stations);
   END_REGION
END_FUNCTION

FUNCTION "Select Buttons: Private: Make Visible / Enable" : Bool   // FC184, SCL
{ S7_Optimized_Access := 'TRUE' }
VERSION : 0.1
   VAR_INPUT
      settings_meta : "Setting Meta Data";
      stations : "Station: All Stations";
   END_VAR
   VAR_TEMP
      ret : Bool;
      enable : Bool;
      is_hmi_station : Bool;
   END_VAR
BEGIN
   REGION "STATIONS ARE HMI STATIONS"
       #is_hmi_station := "Is_HMI_Station"(#stations.stn["Get First Selected Station"(#settings_meta.selected_stations.stns)]);
   END_REGION

